// TIA Portal project "ProjektZaliczenie" (V13) (continued)
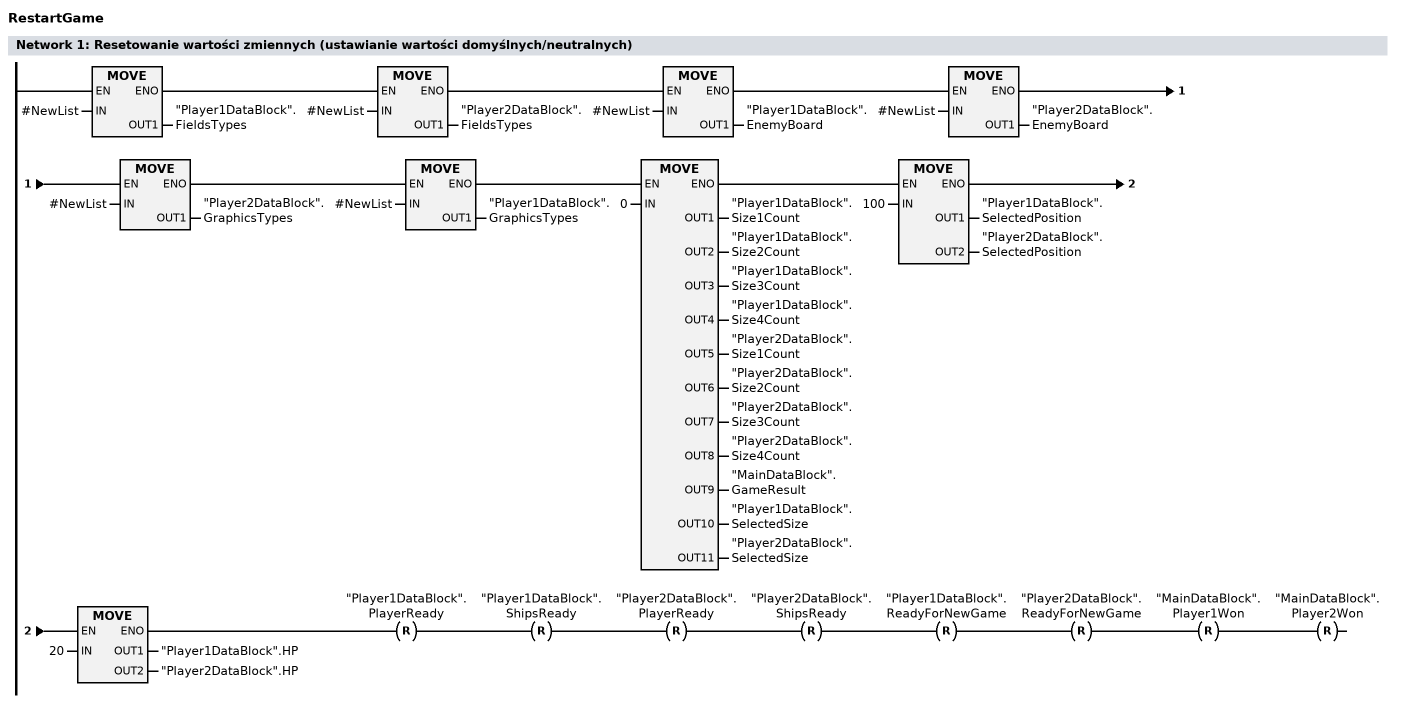
   RUNG wire#powerrail
      { S7_GenerateENO := "TRUE" } Move(in := #NewList, out1 => "Player1DataBlock".FieldsTypes)
      { S7_GenerateENO := "TRUE" } Move(in := #NewList, out1 => "Player2DataBlock".FieldsTypes)
      { S7_GenerateENO := "TRUE" } Move(in := #NewList, out1 => "Player1DataBlock".EnemyBoard)
      { S7_GenerateENO := "TRUE" } Move(in := #NewList, out1 => "Player2DataBlock".EnemyBoard)
      { S7_GenerateENO := "TRUE" } Move(in := #NewList, out1 => "Player2DataBlock".GraphicsTypes)
      { S7_GenerateENO := "TRUE" } Move(in := #NewList, out1 => "Player1DataBlock".GraphicsTypes)
      { S7_GenerateENO := "TRUE" } Move(in := 0, out1 => "Player1DataBlock".Size1Count, out2 => "Player1DataBlock".Size2Count, out3 => "Player1DataBlock".Size3Count, out4 => "Player1DataBlock".Size4Count, out5 => "Player2DataBlock".Size1Count, out6 => "Player2DataBlock".Size2Count, out7 => "Player2DataBlock".Size3Count, out8 => "Player2DataBlock".Size4Count, out9 => "MainDataBlock".GameResult, out10 => "Player1DataBlock".SelectedSize, out11 => "Player2DataBlock".SelectedSize)
      { S7_GenerateENO := "TRUE" } Move(in := 100, out1 => "Player1DataBlock".SelectedPosition, out2 => "Player2DataBlock".SelectedPosition)
      { S7_GenerateENO := "TRUE" } Move(in := 20, out1 => "Player1DataBlock".HP, out2 => "Player2DataBlock".HP)
      R_Coil( "Player1DataBlock".PlayerReady )
      R_Coil( "Player1DataBlock".ShipsReady )
      R_Coil( "Player2DataBlock".PlayerReady )
      R_Coil( "Player2DataBlock".ShipsReady )
      R_Coil( "Player1DataBlock".ReadyForNewGame )
      R_Coil( "Player2DataBlock".ReadyForNewGame )
      R_Coil( "MainDataBlock".Player1Won )
      R_Coil( "MainDataBlock".Player2Won )
   END_RUNG
   // the same network as SCL:
   // ENO of a box is taken as its EN; it also drops when the box reports an error
   "Player1DataBlock".FieldsTypes := #NewList;
   "Player2DataBlock".FieldsTypes := #NewList;
   "Player1DataBlock".EnemyBoard := #NewList;
   "Player2DataBlock".EnemyBoard := #NewList;
   "Player2DataBlock".GraphicsTypes := #NewList;
   "Player1DataBlock".GraphicsTypes := #NewList;
   "Player1DataBlock".Size1Count := 0;
   "Player1DataBlock".Size2Count := 0;
   "Player1DataBlock".Size3Count := 0;
   "Player1DataBlock".Size4Count := 0;
   "Player2DataBlock".Size1Count := 0;
   "Player2DataBlock".Size2Count := 0;
   "Player2DataBlock".Size3Count := 0;
   "Player2DataBlock".Size4Count := 0;
   "MainDataBlock".GameResult := 0;
   "Player1DataBlock".SelectedSize := 0;
   "Player2DataBlock".SelectedSize := 0;
   "Player1DataBlock".SelectedPosition := 100;
   "Player2DataBlock".SelectedPosition := 100;
   "Player1DataBlock".HP := 20;
   "Player2DataBlock".HP := 20;
   "Player1DataBlock".PlayerReady := FALSE;
   "Player1DataBlock".ShipsReady := FALSE;
   "Player2DataBlock".PlayerReady := FALSE;
   "Player2DataBlock".ShipsReady := FALSE;
   "Player1DataBlock".ReadyForNewGame := FALSE;
   "Player2DataBlock".ReadyForNewGame := FALSE;
   "MainDataBlock".Player1Won := FALSE;
   "MainDataBlock".Player2Won := FALSE;
END_REGION
END_FUNCTION_BLOCK

FUNCTION_BLOCK "ResetShips"   // FB5, LAD
TITLE = Resetowanie rozmieszczonych statków
{ S7_Optimized_Access := 'FALSE' }
VERSION : 0.1
BEGIN

REGION Network 1: Ustawianie zmiennych na wartości domyślne/neutralne
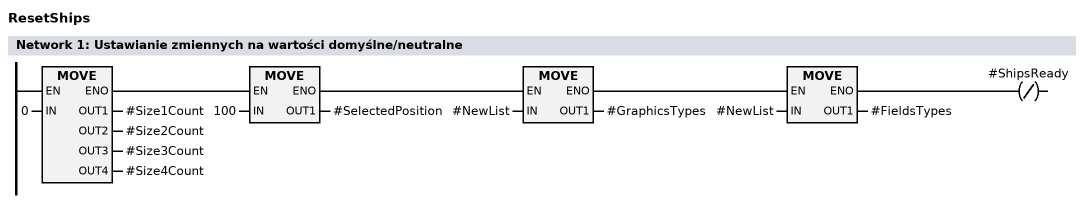
   RUNG wire#powerrail
      { S7_GenerateENO := "TRUE" } Move(in := 0, out1 => #Size1Count, out2 => #Size2Count, out3 => #Size3Count, out4 => #Size4Count)
      { S7_GenerateENO := "TRUE" } Move(in := 100, out1 => #SelectedPosition)
      { S7_GenerateENO := "TRUE" } Move(in := #NewList, out1 => #GraphicsTypes)
      { S7_GenerateENO := "TRUE" } Move(in := #NewList, out1 => #FieldsTypes)
      I_Coil( #ShipsReady )
   END_RUNG
   // the same network as SCL:
   // ENO of a box is taken as its EN; it also drops when the box reports an error
   #Size1Count := 0;
   #Size2Count := 0;
   #Size3Count := 0;
   #Size4Count := 0;
   #SelectedPosition := 100;
   #GraphicsTypes := #NewList;
   #FieldsTypes := #NewList;
   #ShipsReady := NOT TRUE;
END_REGION
END_FUNCTION_BLOCK

FUNCTION "DrawShip" : Void   // FC1, LAD
TITLE = Rysowanie statków
{ S7_Optimized_Access := 'FALSE' }
VERSION : 0.1
// Funkcja odpowiada za rysowanie statkó na planszy (podmienia grafiki na przyciskach)
   VAR_TEMP   // added for the SCL form of the ladder/FBD networks
      _w1 : Bool;
      _w2 : Bool;
      _w3 : Bool;
   END_VAR
BEGIN

REGION Network 1: Setup
   // Ustawianie zmiennych przechowujących informacje o 4 kolejnych polach wertykalnie oraz horyzontalnie
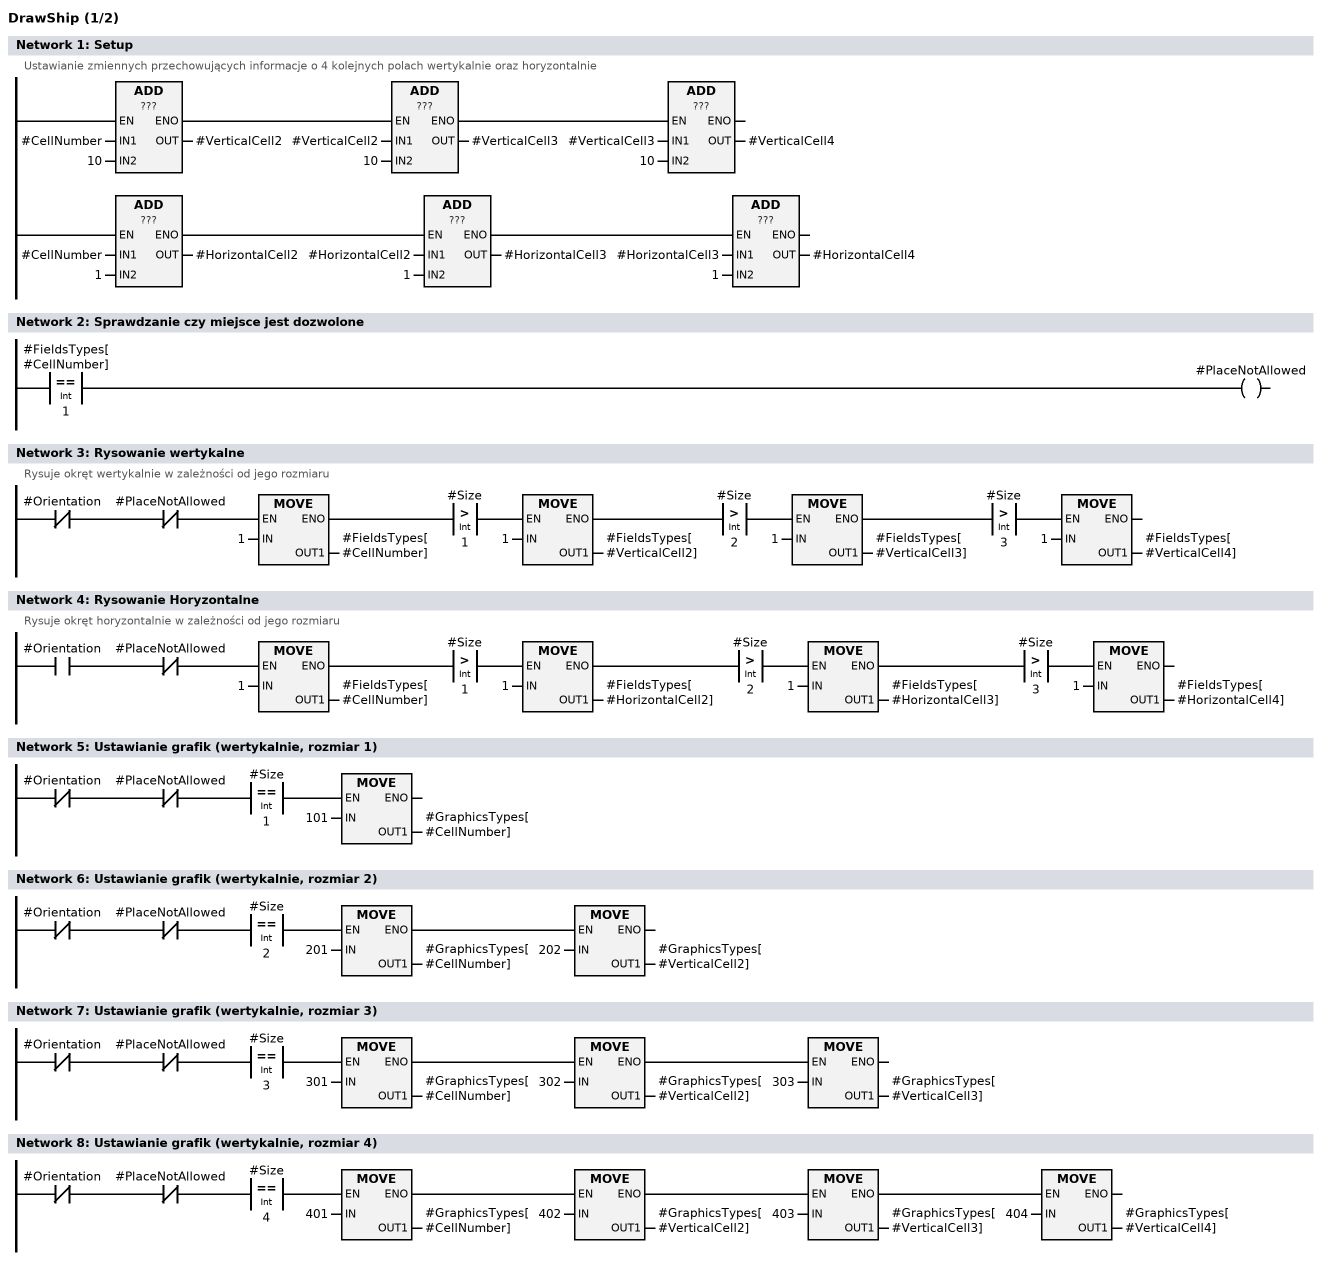
   RUNG wire#powerrail
      { S7_Templates := "SrcType := ???" } Add(in1 := #CellNumber, in2 := 10, out => #VerticalCell2)
      { S7_Templates := "SrcType := ???" } Add(in1 := #VerticalCell2, in2 := 10, out => #VerticalCell3)
      { S7_Templates := "SrcType := ???" } Add(in1 := #VerticalCell3, in2 := 10, out => #VerticalCell4)
   END_RUNG
   RUNG wire#powerrail
      { S7_Templates := "SrcType := ???" } Add(in1 := #CellNumber, in2 := 1, out => #HorizontalCell2)
      { S7_Templates := "SrcType := ???" } Add(in1 := #HorizontalCell2, in2 := 1, out => #HorizontalCell3)
      { S7_Templates := "SrcType := ???" } Add(in1 := #HorizontalCell3, in2 := 1, out => #HorizontalCell4)
   END_RUNG
   // the same network as SCL:
   #VerticalCell2 := #CellNumber + 10;
   #VerticalCell3 := #VerticalCell2 + 10;
   #VerticalCell4 := #VerticalCell3 + 10;
   #HorizontalCell2 := #CellNumber + 1;
   #HorizontalCell3 := #HorizontalCell2 + 1;
   #HorizontalCell4 := #HorizontalCell3 + 1;
END_REGION

REGION Network 2: Sprawdzanie czy miejsce jest dozwolone
   RUNG wire#powerrail
      { S7_Templates := "SrcType := Int" } EQ_Contact(in1 := #FieldsTypes[#CellNumber], in2 := 1)
      Coil( #PlaceNotAllowed )
   END_RUNG
   // the same network as SCL:
   #PlaceNotAllowed := #FieldsTypes[#CellNumber] = 1;
END_REGION

REGION Network 3: Rysowanie wertykalne
   // Rysuje okręt wertykalnie w zależności od jego rozmiaru
   RUNG wire#powerrail
      I_Contact( #Orientation )
      I_Contact( #PlaceNotAllowed )
      Move(in := 1, out1 => #FieldsTypes[#CellNumber])
      { S7_Templates := "SrcType := Int" } GT_Contact(in1 := #Size, in2 := 1)
      Move(in := 1, out1 => #FieldsTypes[#VerticalCell2])
      { S7_Templates := "SrcType := Int" } GT_Contact(in1 := #Size, in2 := 2)
      Move(in := 1, out1 => #FieldsTypes[#VerticalCell3])
      { S7_Templates := "SrcType := Int" } GT_Contact(in1 := #Size, in2 := 3)
      Move(in := 1, out1 => #FieldsTypes[#VerticalCell4])
   END_RUNG
   // the same network as SCL:
   #_w1 := NOT #Orientation AND NOT #PlaceNotAllowed;
   IF #_w1 THEN #FieldsTypes[#CellNumber] := 1; END_IF;
   #_w2 := #_w1 AND (#Size > 1);
   IF #_w2 THEN #FieldsTypes[#VerticalCell2] := 1; END_IF;
   #_w3 := #_w2 AND (#Size > 2);
   IF #_w3 THEN #FieldsTypes[#VerticalCell3] := 1; END_IF;
   IF #_w3 AND (#Size > 3) THEN #FieldsTypes[#VerticalCell4] := 1; END_IF;
END_REGION

REGION Network 4: Rysowanie Horyzontalne
   // Rysuje okręt horyzontalnie w zależności od jego rozmiaru
   RUNG wire#powerrail
      Contact( #Orientation )
      I_Contact( #PlaceNotAllowed )
      Move(in := 1, out1 => #FieldsTypes[#CellNumber])
      { S7_Templates := "SrcType := Int" } GT_Contact(in1 := #Size, in2 := 1)
      Move(in := 1, out1 => #FieldsTypes[#HorizontalCell2])
      { S7_Templates := "SrcType := Int" } GT_Contact(in1 := #Size, in2 := 2)
      Move(in := 1, out1 => #FieldsTypes[#HorizontalCell3])
      { S7_Templates := "SrcType := Int" } GT_Contact(in1 := #Size, in2 := 3)
      Move(in := 1, out1 => #FieldsTypes[#HorizontalCell4])
   END_RUNG
   // the same network as SCL:
   #_w1 := #Orientation AND NOT #PlaceNotAllowed;
   IF #_w1 THEN #FieldsTypes[#CellNumber] := 1; END_IF;
   #_w2 := #_w1 AND (#Size > 1);
   IF #_w2 THEN #FieldsTypes[#HorizontalCell2] := 1; END_IF;
   #_w3 := #_w2 AND (#Size > 2);
   IF #_w3 THEN #FieldsTypes[#HorizontalCell3] := 1; END_IF;
   IF #_w3 AND (#Size > 3) THEN #FieldsTypes[#HorizontalCell4] := 1; END_IF;
END_REGION

REGION Network 5: Ustawianie grafik (wertykalnie, rozmiar 1)
   RUNG wire#powerrail
      I_Contact( #Orientation )
      I_Contact( #PlaceNotAllowed )
      { S7_Templates := "SrcType := Int" } EQ_Contact(in1 := #Size, in2 := 1)
      Move(in := 101, out1 => #GraphicsTypes[#CellNumber])
   END_RUNG
   // the same network as SCL:
   IF NOT #Orientation AND NOT #PlaceNotAllowed AND (#Size = 1) THEN
       #GraphicsTypes[#CellNumber] := 101;
   END_IF;
END_REGION

REGION Network 6: Ustawianie grafik (wertykalnie, rozmiar 2)
   RUNG wire#powerrail
      I_Contact( #Orientation )
      I_Contact( #PlaceNotAllowed )
      { S7_Templates := "SrcType := Int" } EQ_Contact(in1 := #Size, in2 := 2)
      Move(in := 201, out1 => #GraphicsTypes[#CellNumber])
      Move(in := 202, out1 => #GraphicsTypes[#VerticalCell2])
   END_RUNG
   // the same network as SCL:
   IF NOT #Orientation AND NOT #PlaceNotAllowed AND (#Size = 2) THEN
       #GraphicsTypes[#CellNumber] := 201;
       #GraphicsTypes[#VerticalCell2] := 202;
   END_IF;
END_REGION

REGION Network 7: Ustawianie grafik (wertykalnie, rozmiar 3)
   RUNG wire#powerrail
      I_Contact( #Orientation )
      I_Contact( #PlaceNotAllowed )
      { S7_Templates := "SrcType := Int" } EQ_Contact(in1 := #Size, in2 := 3)
      Move(in := 301, out1 => #GraphicsTypes[#CellNumber])
      Move(in := 302, out1 => #GraphicsTypes[#VerticalCell2])
      Move(in := 303, out1 => #GraphicsTypes[#VerticalCell3])
   END_RUNG
   // the same network as SCL:
   IF NOT #Orientation AND NOT #PlaceNotAllowed AND (#Size = 3) THEN
       #GraphicsTypes[#CellNumber] := 301;
       #GraphicsTypes[#VerticalCell2] := 302;
       #GraphicsTypes[#VerticalCell3] := 303;
   END_IF;
END_REGION

REGION Network 8: Ustawianie grafik (wertykalnie, rozmiar 4)
   RUNG wire#powerrail
      I_Contact( #Orientation )
      I_Contact( #PlaceNotAllowed )
      { S7_Templates := "SrcType := Int" } EQ_Contact(in1 := #Size, in2 := 4)
      Move(in := 401, out1 => #GraphicsTypes[#CellNumber])
      Move(in := 402, out1 => #GraphicsTypes[#VerticalCell2])
      Move(in := 403, out1 => #GraphicsTypes[#VerticalCell3])
      Move(in := 404, out1 => #GraphicsTypes[#VerticalCell4])
   END_RUNG
   // the same network as SCL:
   IF NOT #Orientation AND NOT #PlaceNotAllowed AND (#Size = 4) THEN
       #GraphicsTypes[#CellNumber] := 401;
       #GraphicsTypes[#VerticalCell2] := 402;
       #GraphicsTypes[#VerticalCell3] := 403;
       #GraphicsTypes[#VerticalCell4] := 404;
   END_IF;
END_REGION

REGION Network 9: Ustawianie grafik (horyzontalnie, rozmiar 1)
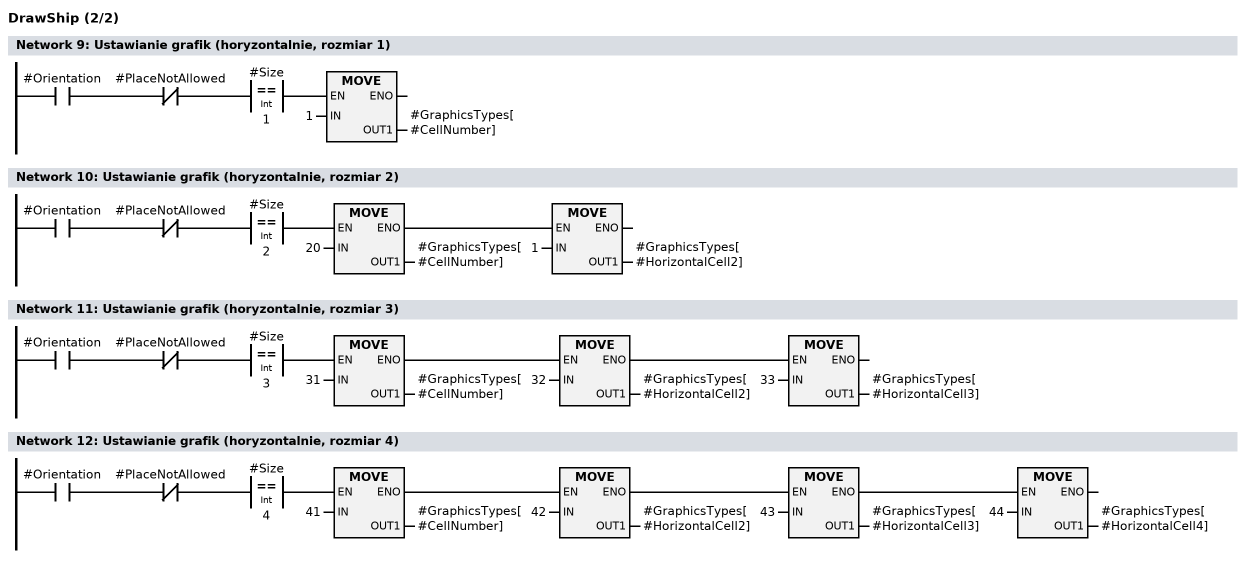
   RUNG wire#powerrail
      Contact( #Orientation )
      I_Contact( #PlaceNotAllowed )
      { S7_Templates := "SrcType := Int" } EQ_Contact(in1 := #Size, in2 := 1)
      Move(in := 1, out1 => #GraphicsTypes[#CellNumber])
   END_RUNG
   // the same network as SCL:
   IF #Orientation AND NOT #PlaceNotAllowed AND (#Size = 1) THEN #GraphicsTypes[#CellNumber] := 1; END_IF;
END_REGION

REGION Network 10: Ustawianie grafik (horyzontalnie, rozmiar 2)
   RUNG wire#powerrail
      Contact( #Orientation )
      I_Contact( #PlaceNotAllowed )
      { S7_Templates := "SrcType := Int" } EQ_Contact(in1 := #Size, in2 := 2)
      Move(in := 20, out1 => #GraphicsTypes[#CellNumber])
      Move(in := 1, out1 => #GraphicsTypes[#HorizontalCell2])
   END_RUNG
   // the same network as SCL:
   IF #Orientation AND NOT #PlaceNotAllowed AND (#Size = 2) THEN
       #GraphicsTypes[#CellNumber] := 20;
       #GraphicsTypes[#HorizontalCell2] := 1;
   END_IF;
END_REGION

REGION Network 11: Ustawianie grafik (horyzontalnie, rozmiar 3)
   RUNG wire#powerrail
      Contact( #Orientation )
      I_Contact( #PlaceNotAllowed )
      { S7_Templates := "SrcType := Int" } EQ_Contact(in1 := #Size, in2 := 3)
      Move(in := 31, out1 => #GraphicsTypes[#CellNumber])
      Move(in := 32, out1 => #GraphicsTypes[#HorizontalCell2])
      Move(in := 33, out1 => #GraphicsTypes[#HorizontalCell3])
   END_RUNG
   // the same network as SCL:
   IF #Orientation AND NOT #PlaceNotAllowed AND (#Size = 3) THEN
       #GraphicsTypes[#CellNumber] := 31;
       #GraphicsTypes[#HorizontalCell2] := 32;
       #GraphicsTypes[#HorizontalCell3] := 33;
   END_IF;
END_REGION

REGION Network 12: Ustawianie grafik (horyzontalnie, rozmiar 4)
   RUNG wire#powerrail
      Contact( #Orientation )
      I_Contact( #PlaceNotAllowed )
      { S7_Templates := "SrcType := Int" } EQ_Contact(in1 := #Size, in2 := 4)
      Move(in := 41, out1 => #GraphicsTypes[#CellNumber])
      Move(in := 42, out1 => #GraphicsTypes[#HorizontalCell2])
      Move(in := 43, out1 => #GraphicsTypes[#HorizontalCell3])
      Move(in := 44, out1 => #GraphicsTypes[#HorizontalCell4])
   END_RUNG
   // the same network as SCL:
   IF #Orientation AND NOT #PlaceNotAllowed AND (#Size = 4) THEN
       #GraphicsTypes[#CellNumber] := 41;
       #GraphicsTypes[#HorizontalCell2] := 42;
       #GraphicsTypes[#HorizontalCell3] := 43;
       #GraphicsTypes[#HorizontalCell4] := 44;
   END_IF;
END_REGION
END_FUNCTION

FUNCTION "CheckPosition" : Void   // FC2, SCL
{ S7_Optimized_Access := 'FALSE' }
VERSION : 0.1
BEGIN
   IF #Orientation THEN // Orientacja horyzontalna
       IF (#CellNumber MOD 10) = 0 THEN // Lewa granica mapy (Nie potrzeba sprawdzać komórki na lewo)
           #Start := #CellNumber;
       ELSE
           #Start := #CellNumber - 1;
       END_IF;

       IF ((#CellNumber + #Size - 1) MOD 10) = 9 THEN // Prawa granica mapy (Nie potrzeba sprawdzać komórki na prawo)
           #End := #CellNumber + #Size - 1;
       ELSE
           #End := #CellNumber + #Size;
       END_IF;

       IF #Start MOD 10 > #End MOD 10 THEN // Część statku znajduje się już w następnym rzędzie (Statek jest zbyt duży)
           #PositionNotAllowed := 1;
       ELSE
           FOR #i := #Start TO #End DO // Pętla sprawdzająca czy okręt nie styka się z pozostałymi statkami 

               IF #FieldsTypes[#i] = 1 THEN
                   #PositionNotAllowed := 1;
                   EXIT;
               END_IF;

               IF #Start - 10 >= 0 THEN // Nie potrzeba sprawdzać komórek powyżej (statek ustawiony jest przy górnej granicy mapy)
                   IF #FieldsTypes[#i - 10] = 1 THEN
                       #PositionNotAllowed := 1;
                       EXIT;
                   END_IF;

               END_IF;

               IF #Start + 10 <= 99 THEN // Nie potrzeba sprawdzać komórek poniżej (statek ustawiony jest przy dolnej granicy mapy)
                   IF #FieldsTypes[#i + 10] = 1 THEN
                       #PositionNotAllowed := 1;
                       EXIT;
                   END_IF;

               END_IF;


           END_FOR;

       END_IF;

   ELSE // Orientacja wertykalna
       IF #CellNumber  < 10 THEN // Nie potrzeba sprawdzać komórek powyżej (górna granica mapy)
           #Start := #CellNumber;
       ELSE
           #Start := #CellNumber - 10;
       END_IF;

       IF (#CellNumber + ((#Size - 1) * 10)) <= 99 AND (#CellNumber + ((#Size - 1) * 10)) >= 90 THEN // Bottom map border (We do not need to check cell below)
           #End := #CellNumber + ((#Size - 1) * 10);
       ELSE
           #End := #CellNumber + (#Size * 10);
       END_IF;

       IF #End > 99 THEN // Statek jest za duży
           #PositionNotAllowed := 1;
       ELSE
           FOR #i := #Start TO #End BY 10 DO // Pętla sprawdzająca czy okręt nie styka się z pozostałymi statkami 

               IF #FieldsTypes[#i] = 1 THEN
                   #PositionNotAllowed := 1;
                   EXIT;
               END_IF;

               IF (#i MOD 10) > 0 THEN // Nie potrzeba sprawdzać komórek po lewej (statek znajduje się przy lewej granicy mapy)
                   IF #FieldsTypes[#i - 1] = 1 THEN
                       #PositionNotAllowed := 1;
                       EXIT;
                   END_IF;
               END_IF;

               IF (#i MOD 10) < 9 THEN // Nie potrzeba sprawdzać komórek po prawej (statek znadjduje się przy prawej granicy mapy)
                   IF #FieldsTypes[#i + 1] = 1 THEN
                       #PositionNotAllowed := 1;
                       EXIT;
                   END_IF;
               END_IF;

           END_FOR;

       END_IF;



   END_IF;
END_FUNCTION

FUNCTION "CountShips" : Void   // FC3, LAD
TITLE = Liczenie okrętów
{ S7_Optimized_Access := 'FALSE' }
VERSION : 0.1
// Funkcja zliczająca okręty określonych rozmiarów oraz informująca o rozmieszczeniu wszystkich okrętów
   VAR_TEMP   // added for the SCL form of the ladder/FBD networks
      _w1 : Bool;
      _w2 : Bool;
      _w3 : Bool;
      _w4 : Bool;
   END_VAR
BEGIN

REGION Network 1: Wystawianie danych wejściowych bezpośrednio na wyjście
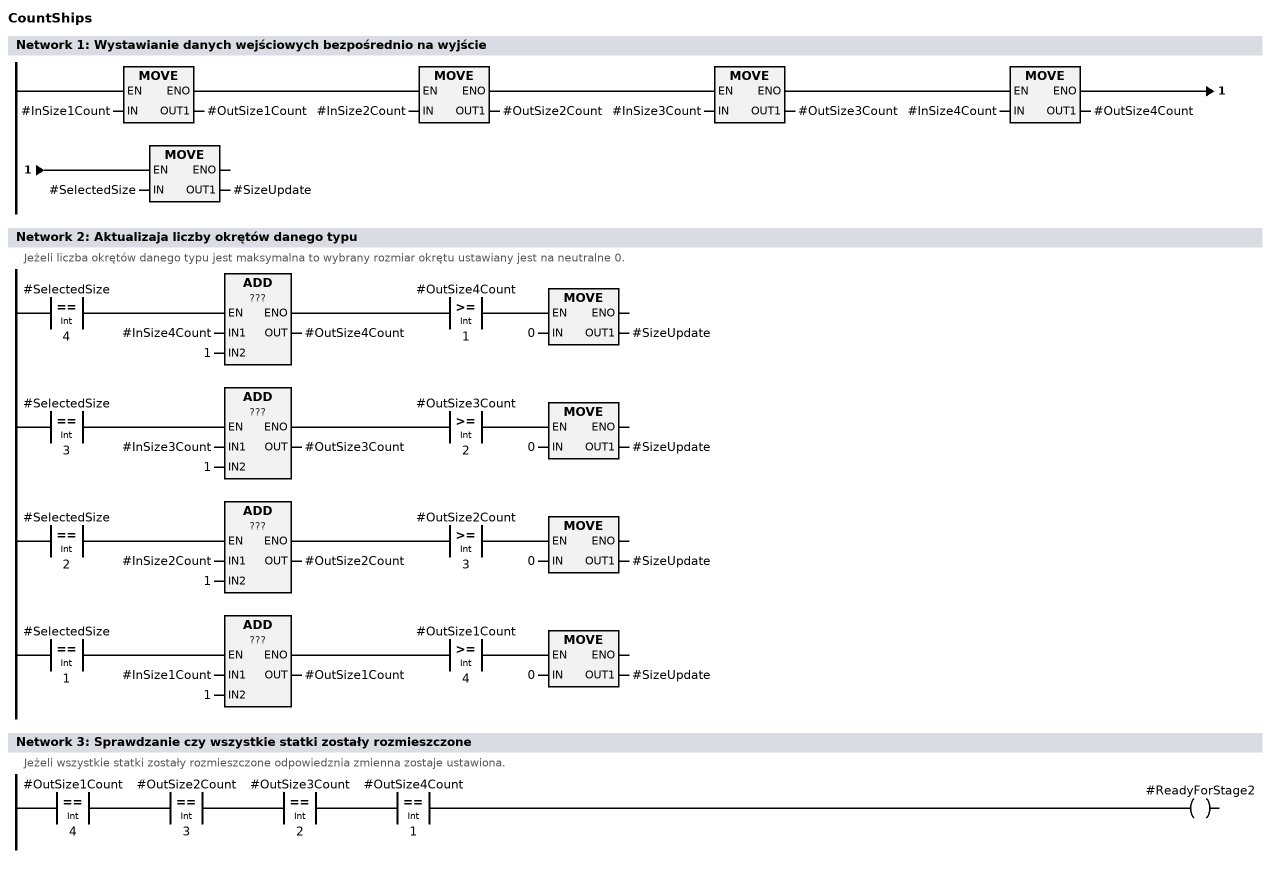
   RUNG wire#powerrail
      Move(in := #InSize1Count, out1 => #OutSize1Count)
      Move(in := #InSize2Count, out1 => #OutSize2Count)
      Move(in := #InSize3Count, out1 => #OutSize3Count)
      Move(in := #InSize4Count, out1 => #OutSize4Count)
      Move(in := #SelectedSize, out1 => #SizeUpdate)
   END_RUNG
   // the same network as SCL:
   #OutSize1Count := #InSize1Count;
   #OutSize2Count := #InSize2Count;
   #OutSize3Count := #InSize3Count;
   #OutSize4Count := #InSize4Count;
   #SizeUpdate := #SelectedSize;
END_REGION

REGION Network 2: Aktualizaja liczby okrętów danego typu
   // Jeżeli liczba okrętów danego typu jest maksymalna to wybrany rozmiar okrętu ustawiany jest na neutralne 0.
   RUNG wire#powerrail
      { S7_Templates := "SrcType := Int" } EQ_Contact(in1 := #SelectedSize, in2 := 4)
      { S7_Templates := "SrcType := ???" } Add(in1 := #InSize4Count, in2 := 1, out => #OutSize4Count)
      { S7_Templates := "SrcType := Int" } GE_Contact(in1 := #OutSize4Count, in2 := 1)
      Move(in := 0, out1 => #SizeUpdate)
   END_RUNG
   RUNG wire#powerrail
      { S7_Templates := "SrcType := Int" } EQ_Contact(in1 := #SelectedSize, in2 := 3)
      { S7_Templates := "SrcType := ???" } Add(in1 := #InSize3Count, in2 := 1, out => #OutSize3Count)
      { S7_Templates := "SrcType := Int" } GE_Contact(in1 := #OutSize3Count, in2 := 2)
      Move(in := 0, out1 => #SizeUpdate)
   END_RUNG
   RUNG wire#powerrail
      { S7_Templates := "SrcType := Int" } EQ_Contact(in1 := #SelectedSize, in2 := 2)
      { S7_Templates := "SrcType := ???" } Add(in1 := #InSize2Count, in2 := 1, out => #OutSize2Count)
      { S7_Templates := "SrcType := Int" } GE_Contact(in1 := #OutSize2Count, in2 := 3)
      Move(in := 0, out1 => #SizeUpdate)
   END_RUNG
   RUNG wire#powerrail
      { S7_Templates := "SrcType := Int" } EQ_Contact(in1 := #SelectedSize, in2 := 1)
      { S7_Templates := "SrcType := ???" } Add(in1 := #InSize1Count, in2 := 1, out => #OutSize1Count)
      { S7_Templates := "SrcType := Int" } GE_Contact(in1 := #OutSize1Count, in2 := 4)
      Move(in := 0, out1 => #SizeUpdate)
   END_RUNG
   // the same network as SCL:
   #_w1 := #SelectedSize = 4;
   IF #_w1 THEN #OutSize4Count := #InSize4Count + 1; END_IF;
   IF #_w1 AND (#OutSize4Count >= 1) THEN #SizeUpdate := 0; END_IF;
   #_w2 := #SelectedSize = 3;
   IF #_w2 THEN #OutSize3Count := #InSize3Count + 1; END_IF;
   IF #_w2 AND (#OutSize3Count >= 2) THEN #SizeUpdate := 0; END_IF;
   #_w3 := #SelectedSize = 2;
   IF #_w3 THEN #OutSize2Count := #InSize2Count + 1; END_IF;
   IF #_w3 AND (#OutSize2Count >= 3) THEN #SizeUpdate := 0; END_IF;
   #_w4 := #SelectedSize = 1;
   IF #_w4 THEN #OutSize1Count := #InSize1Count + 1; END_IF;
   IF #_w4 AND (#OutSize1Count >= 4) THEN #SizeUpdate := 0; END_IF;
END_REGION

REGION Network 3: Sprawdzanie czy wszystkie statki zostały rozmieszczone
   // Jeżeli wszystkie statki zostały rozmieszczone odpowiedznia zmienna zostaje ustawiona.
   RUNG wire#powerrail
      { S7_Templates := "SrcType := Int" } EQ_Contact(in1 := #OutSize1Count, in2 := 4)
      { S7_Templates := "SrcType := Int" } EQ_Contact(in1 := #OutSize2Count, in2 := 3)
      { S7_Templates := "SrcType := Int" } EQ_Contact(in1 := #OutSize3Count, in2 := 2)
      { S7_Templates := "SrcType := Int" } EQ_Contact(in1 := #OutSize4Count, in2 := 1)
      Coil( #ReadyForStage2 )
   END_RUNG
   // the same network as SCL:
   #ReadyForStage2 := (#OutSize1Count = 4) AND (#OutSize2Count = 3) AND (#OutSize3Count = 2) AND (#OutSize4Count = 1);
END_REGION
END_FUNCTION

FUNCTION "ChangeScreen" : Void   // FC5, LAD
TITLE = Zmiana ekranu
{ S7_Optimized_Access := 'FALSE' }
VERSION : 0.1
// Funkcja wysyła do paneli HMI żądanie zmiany ekranu
BEGIN

REGION Network 1: Ekran 1
   // 51 - zmień ekran
   // ScreenNumber - nr ekranu
   // 0 - bez znaczenia
   // 0 - bez znaczenia
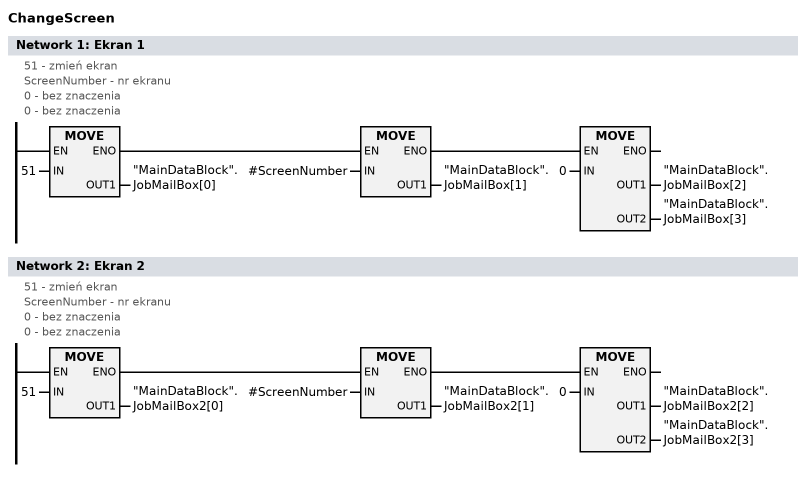
   RUNG wire#powerrail
      { S7_GenerateENO := "TRUE" } Move(in := 51, out1 => "MainDataBlock".JobMailBox[0])
      { S7_GenerateENO := "TRUE" } Move(in := #ScreenNumber, out1 => "MainDataBlock".JobMailBox[1])
      { S7_GenerateENO := "TRUE" } Move(in := 0, out1 => "MainDataBlock".JobMailBox[2], out2 => "MainDataBlock".JobMailBox[3])
   END_RUNG
   // the same network as SCL:
   // ENO of a box is taken as its EN; it also drops when the box reports an error
   "MainDataBlock".JobMailBox[0] := 51;
   "MainDataBlock".JobMailBox[1] := #ScreenNumber;
   "MainDataBlock".JobMailBox[2] := 0;
   "MainDataBlock".JobMailBox[3] := 0;
END_REGION

REGION Network 2: Ekran 2
   // 51 - zmień ekran
   // ScreenNumber - nr ekranu
   // 0 - bez znaczenia
   // 0 - bez znaczenia
   RUNG wire#powerrail
      { S7_GenerateENO := "TRUE" } Move(in := 51, out1 => "MainDataBlock".JobMailBox2[0])
      { S7_GenerateENO := "TRUE" } Move(in := #ScreenNumber, out1 => "MainDataBlock".JobMailBox2[1])
      { S7_GenerateENO := "TRUE" } Move(in := 0, out1 => "MainDataBlock".JobMailBox2[2], out2 => "MainDataBlock".JobMailBox2[3])
   END_RUNG
   // the same network as SCL:
   // ENO of a box is taken as its EN; it also drops when the box reports an error
   "MainDataBlock".JobMailBox2[0] := 51;
   "MainDataBlock".JobMailBox2[1] := #ScreenNumber;
   "MainDataBlock".JobMailBox2[2] := 0;
   "MainDataBlock".JobMailBox2[3] := 0;
END_REGION
END_FUNCTION

FUNCTION "CheckHit" : Void   // FC6, LAD
TITLE = Sprawdzanie trafienia
{ S7_Optimized_Access := 'FALSE' }
VERSION : 0.1
// Funkcja sprawdza pole wybrane przez gracza pod kątem obecności wrogiego statku oraz aktualizuje wybrane pole (pudło/trafienie).
   VAR_TEMP   // added for the SCL form of the ladder/FBD networks
      _w1 : Bool;
   END_VAR
BEGIN

REGION Network 1: Pudło
   // Informacja o braku trafienia (zmienna HIT) oraz aktualizacja pól (zmiana grafik oraz typów).
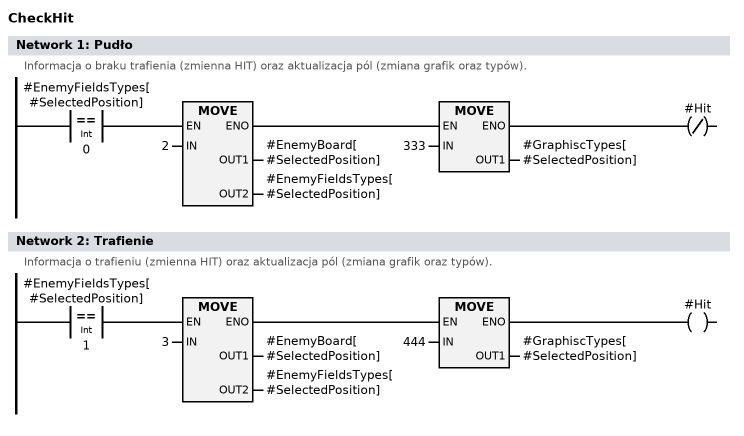
   RUNG wire#powerrail
      { S7_Templates := "SrcType := Int" } EQ_Contact(in1 := #EnemyFieldsTypes[#SelectedPosition], in2 := 0)
      { S7_GenerateENO := "TRUE" } Move(in := 2, out1 => #EnemyBoard[#SelectedPosition], out2 => #EnemyFieldsTypes[#SelectedPosition])
      { S7_GenerateENO := "TRUE" } Move(in := 333, out1 => #GraphiscTypes[#SelectedPosition])
      I_Coil( #Hit )
   END_RUNG
   // the same network as SCL:
   // ENO of a box is taken as its EN; it also drops when the box reports an error
   #_w1 := #EnemyFieldsTypes[#SelectedPosition] = 0;
   IF #_w1 THEN
       #EnemyBoard[#SelectedPosition] := 2;
       #EnemyFieldsTypes[#SelectedPosition] := 2;
       #GraphiscTypes[#SelectedPosition] := 333;
   END_IF;
   #Hit := NOT #_w1;
END_REGION

REGION Network 2: Trafienie
   // Informacja o trafieniu (zmienna HIT) oraz aktualizacja pól (zmiana grafik oraz typów).
   RUNG wire#powerrail
      { S7_Templates := "SrcType := Int" } EQ_Contact(in1 := #EnemyFieldsTypes[#SelectedPosition], in2 := 1)
      { S7_GenerateENO := "TRUE" } Move(in := 3, out1 => #EnemyBoard[#SelectedPosition], out2 => #EnemyFieldsTypes[#SelectedPosition])
      { S7_GenerateENO := "TRUE" } Move(in := 444, out1 => #GraphiscTypes[#SelectedPosition])
      Coil( #Hit )
   END_RUNG
   // the same network as SCL:
   // ENO of a box is taken as its EN; it also drops when the box reports an error
   #_w1 := #EnemyFieldsTypes[#SelectedPosition] = 1;
   IF #_w1 THEN
       #EnemyBoard[#SelectedPosition] := 3;
       #EnemyFieldsTypes[#SelectedPosition] := 3;
       #GraphiscTypes[#SelectedPosition] := 444;
   END_IF;
   #Hit := #_w1;
END_REGION
END_FUNCTION

FUNCTION "CheckWin" : Void   // FC7, LAD
TITLE = Sprawdzanie zakończenia gry
{ S7_Optimized_Access := 'FALSE' }
VERSION : 0.1
// Funkcja sprawdza czy któryś z graczy nie utracił wszystkich punktów HP.
BEGIN

REGION Network 1: Gracz 1
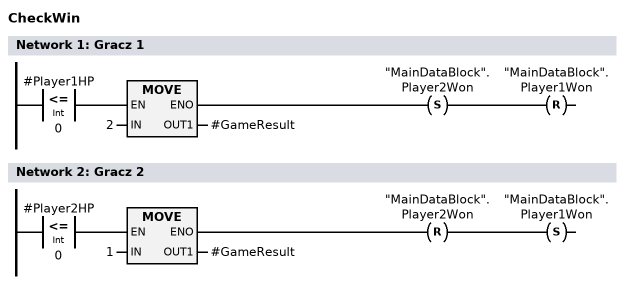
   RUNG wire#powerrail
      { S7_Templates := "SrcType := Int" } LE_Contact(in1 := #Player1HP, in2 := 0)
      { S7_GenerateENO := "TRUE" } Move(in := 2, out1 => #GameResult)
      S_Coil( "MainDataBlock".Player2Won )
      R_Coil( "MainDataBlock".Player1Won )
   END_RUNG
   // the same network as SCL:
   // ENO of a box is taken as its EN; it also drops when the box reports an error
   IF #Player1HP <= 0 THEN
       #GameResult := 2;
       "MainDataBlock".Player2Won := TRUE;
       "MainDataBlock".Player1Won := FALSE;
   END_IF;
END_REGION

REGION Network 2: Gracz 2
   RUNG wire#powerrail
      { S7_Templates := "SrcType := Int" } LE_Contact(in1 := #Player2HP, in2 := 0)
      { S7_GenerateENO := "TRUE" } Move(in := 1, out1 => #GameResult)
      R_Coil( "MainDataBlock".Player2Won )
      S_Coil( "MainDataBlock".Player1Won )
   END_RUNG
   // the same network as SCL:
   // ENO of a box is taken as its EN; it also drops when the box reports an error
   IF #Player2HP <= 0 THEN
       #GameResult := 1;
       "MainDataBlock".Player2Won := FALSE;
       "MainDataBlock".Player1Won := TRUE;
   END_IF;
END_REGION
END_FUNCTION

ORGANIZATION_BLOCK "Main"   // OB1, LAD, ProgramCycle
TITLE = Główny blok programu
{ S7_Optimized_Access := 'FALSE' }
VERSION : 0.1
BEGIN

REGION Network 1: Etap 1
   // Rozmieszczanie statków
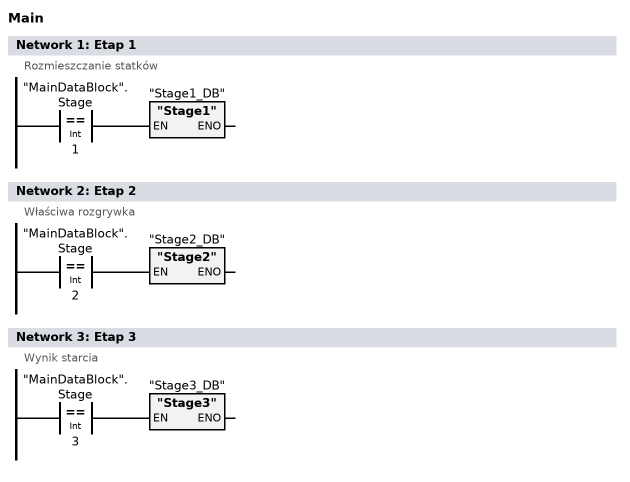
   RUNG wire#powerrail
      { S7_Templates := "SrcType := Int" } EQ_Contact(in1 := "MainDataBlock".Stage, in2 := 1)
      "Stage1_DB"()
   END_RUNG
   // the same network as SCL:
   IF "MainDataBlock".Stage = 1 THEN
       "Stage1_DB"();   // "Stage1"
   END_IF;
END_REGION

REGION Network 2: Etap 2
   // Właściwa rozgrywka
   RUNG wire#powerrail
      { S7_Templates := "SrcType := Int" } EQ_Contact(in1 := "MainDataBlock".Stage, in2 := 2)
      "Stage2_DB"()
   END_RUNG
   // the same network as SCL:
   IF "MainDataBlock".Stage = 2 THEN
       "Stage2_DB"();   // "Stage2"
   END_IF;
END_REGION

REGION Network 3: Etap 3
   // Wynik starcia
   RUNG wire#powerrail
      { S7_Templates := "SrcType := Int" } EQ_Contact(in1 := "MainDataBlock".Stage, in2 := 3)
      "Stage3_DB"()
   END_RUNG
   // the same network as SCL:
   IF "MainDataBlock".Stage = 3 THEN
       "Stage3_DB"();   // "Stage3"
   END_IF;
END_REGION
END_ORGANIZATION_BLOCK

(* ===== HMI "HMI_RT_1" =====
connection "HMI_Connection_1": ETHERNET, SMART_S7_1200_OMS
